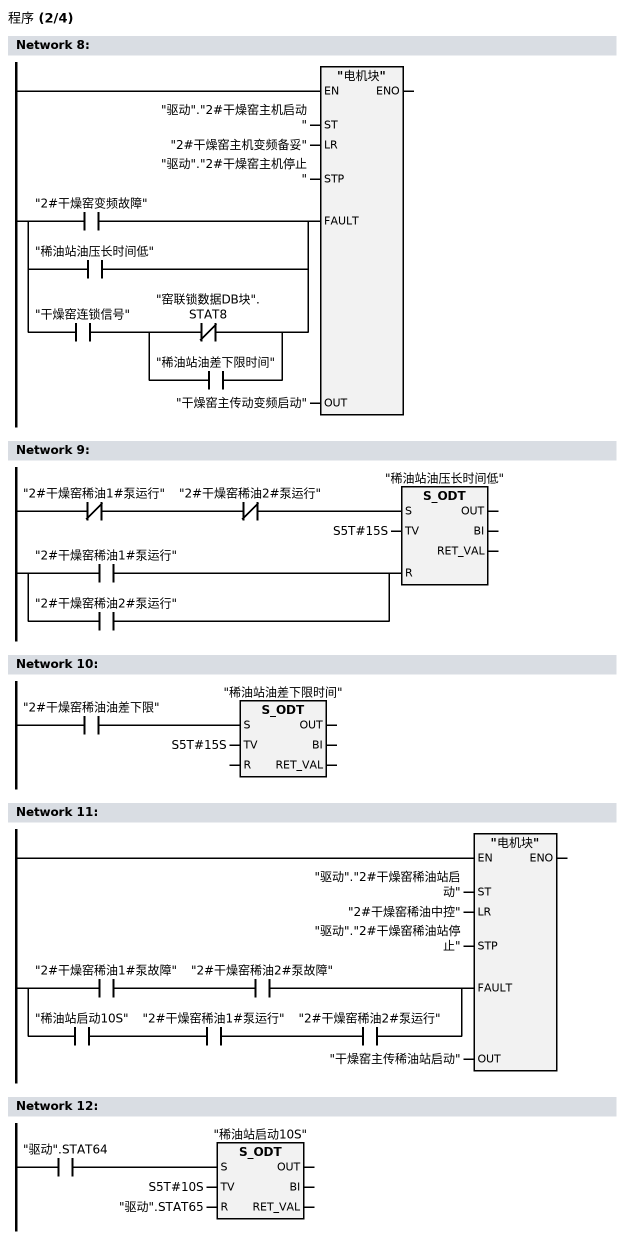
   RUNG wire#powerrail
      "电机块"(FAULT := wire#w2, ST := "驱动"."2#干燥窑主机启动", LR := "2#干燥窑主机变频备妥", STP := "驱动"."2#干燥窑主机停止", OUT := "干燥窑主传动变频启动")
   END_RUNG
   RUNG wire#powerrail
      Contact( "2#干燥窑变频故障" )
   END_RUNG wire#w2
   RUNG wire#powerrail
      Contact( "稀油站油压长时间低" )
   END_RUNG wire#w2
   RUNG wire#powerrail
      Contact( "干燥窑连锁信号" )
      wire#w1
      I_Contact( "窑联锁数据DB块".STAT8 )
   END_RUNG wire#w2
   RUNG wire#w1
      Contact( "稀油站油差下限时间" )
   END_RUNG wire#w2
   // the same network as SCL:
   "电机块"(ST := "驱动"."2#干燥窑主机启动",
         LR := "2#干燥窑主机变频备妥",
         STP := "驱动"."2#干燥窑主机停止",
         FAULT := "2#干燥窑变频故障" OR "稀油站油压长时间低" OR ("干燥窑连锁信号" AND (NOT "窑联锁数据DB块".STAT8 OR "稀油站油差下限时间")),
         OUT := "干燥窑主传动变频启动");
END_REGION

REGION Network 9
   RUNG wire#powerrail
      I_Contact( "2#干燥窑稀油1#泵运行" )
      I_Contact( "2#干燥窑稀油2#泵运行" )
      S_ODT(T_NO := "稀油站油压长时间低", TV := S5T#15S, R := wire#w1, BI =>, RET_VAL =>)
   END_RUNG
   RUNG wire#powerrail
      Contact( "2#干燥窑稀油1#泵运行" )
   END_RUNG wire#w1
   RUNG wire#powerrail
      Contact( "2#干燥窑稀油2#泵运行" )
   END_RUNG wire#w1
   // the same network as SCL:
   #_s5time1 := S_ODT(T_NO := "稀油站油压长时间低",
                      TV := S5T#15S,
                      R := "2#干燥窑稀油1#泵运行" OR "2#干燥窑稀油2#泵运行",
                      S := NOT "2#干燥窑稀油1#泵运行" AND NOT "2#干燥窑稀油2#泵运行");
END_REGION

REGION Network 10
   RUNG wire#powerrail
      Contact( "2#干燥窑稀油油差下限" )
      S_ODT(T_NO := "稀油站油差下限时间", TV := S5T#15S, R :=, BI =>, RET_VAL =>)
   END_RUNG
   // the same network as SCL:
   #_s5time1 := S_ODT(T_NO := "稀油站油差下限时间", TV := S5T#15S, S := "2#干燥窑稀油油差下限");
END_REGION

REGION Network 11
   RUNG wire#powerrail
      "电机块"(FAULT := wire#w1, ST := "驱动"."2#干燥窑稀油站启动", LR := "2#干燥窑稀油中控", STP := "驱动"."2#干燥窑稀油站停止", OUT := "干燥窑主传稀油站启动")
   END_RUNG
   RUNG wire#powerrail
      Contact( "2#干燥窑稀油1#泵故障" )
      Contact( "2#干燥窑稀油2#泵故障" )
   END_RUNG wire#w1
   RUNG wire#powerrail
      Contact( "稀油站启动10S" )
      Contact( "2#干燥窑稀油1#泵运行" )
      Contact( "2#干燥窑稀油2#泵运行" )
   END_RUNG wire#w1
   // the same network as SCL:
   "电机块"(ST := "驱动"."2#干燥窑稀油站启动",
         LR := "2#干燥窑稀油中控",
         STP := "驱动"."2#干燥窑稀油站停止",
         FAULT := ("2#干燥窑稀油1#泵故障" AND "2#干燥窑稀油2#泵故障") OR ("稀油站启动10S" AND "2#干燥窑稀油1#泵运行" AND "2#干燥窑稀油2#泵运行"),
         OUT := "干燥窑主传稀油站启动");
END_REGION

REGION Network 12
   RUNG wire#powerrail
      Contact( "驱动".STAT64 )
      S_ODT(T_NO := "稀油站启动10S", TV := S5T#10S, R := "驱动".STAT65, BI =>, RET_VAL =>)
   END_RUNG
   // the same network as SCL:
   #_s5time1 := S_ODT(T_NO := "稀油站启动10S", S := "驱动".STAT64, TV := S5T#10S, R := "驱动".STAT65);
END_REGION

REGION Network 13
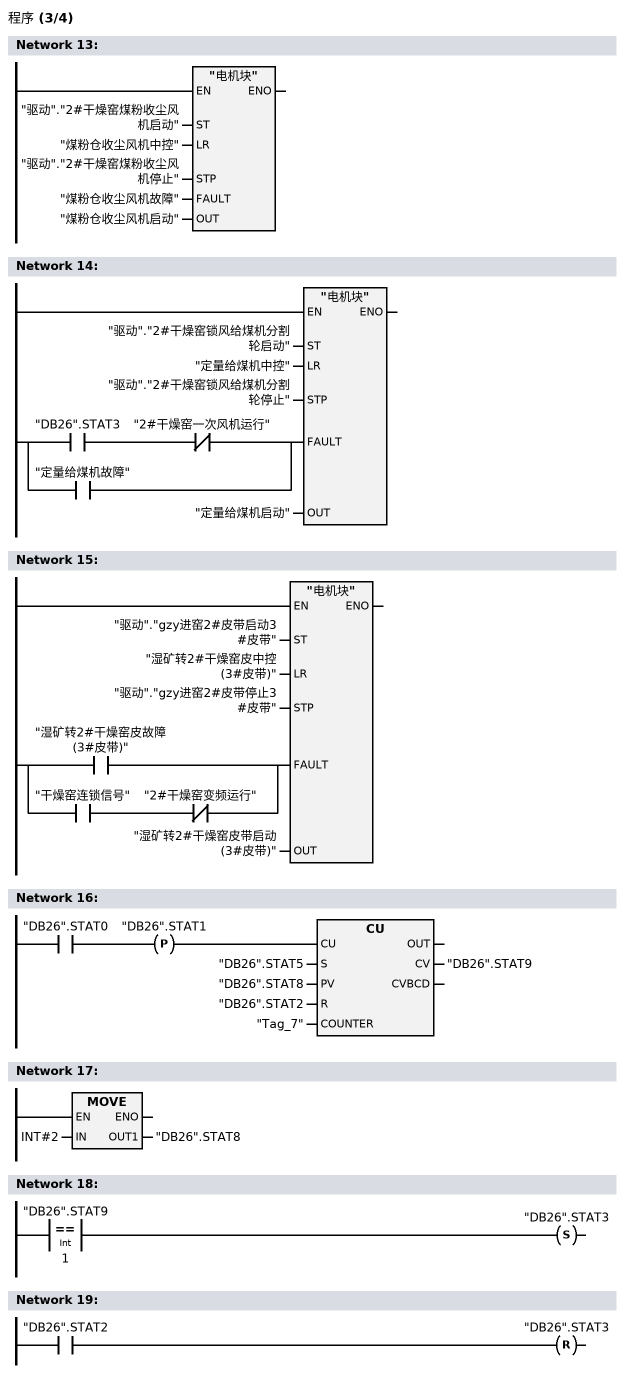
   RUNG wire#powerrail
      "电机块"(ST := "驱动"."2#干燥窑煤粉收尘风机启动", LR := "煤粉仓收尘风机中控", STP := "驱动"."2#干燥窑煤粉收尘风机停止", FAULT := "煤粉仓收尘风机故障", OUT := "煤粉仓收尘风机启动")
   END_RUNG
   // the same network as SCL:
   "电机块"(ST := "驱动"."2#干燥窑煤粉收尘风机启动",
         LR := "煤粉仓收尘风机中控",
         STP := "驱动"."2#干燥窑煤粉收尘风机停止",
         FAULT := "煤粉仓收尘风机故障",
         OUT := "煤粉仓收尘风机启动");
END_REGION

REGION Network 14
   RUNG wire#powerrail
      "电机块"(FAULT := wire#w1, ST := "驱动"."2#干燥窑锁风给煤机分割轮启动", LR := "定量给煤机中控", STP := "驱动"."2#干燥窑锁风给煤机分割轮停止", OUT := "定量给煤机启动")
   END_RUNG
   RUNG wire#powerrail
      Contact( "DB26".STAT3 )
      I_Contact( "2#干燥窑一次风机运行" )
   END_RUNG wire#w1
   RUNG wire#powerrail
      Contact( "定量给煤机故障" )
   END_RUNG wire#w1
   // the same network as SCL:
   "电机块"(ST := "驱动"."2#干燥窑锁风给煤机分割轮启动",
         LR := "定量给煤机中控",
         STP := "驱动"."2#干燥窑锁风给煤机分割轮停止",
         FAULT := ("DB26".STAT3 AND NOT "2#干燥窑一次风机运行") OR "定量给煤机故障",
         OUT := "定量给煤机启动");
END_REGION

REGION Network 15
   RUNG wire#powerrail
      "电机块"(FAULT := wire#w1, ST := "驱动"."gzy进窑2#皮带启动3#皮带", LR := "湿矿转2#干燥窑皮中控  (3#皮带)", STP := "驱动"."gzy进窑2#皮带停止3#皮带", OUT := "湿矿转2#干燥窑皮带启动  (3#皮带)")
   END_RUNG
   RUNG wire#powerrail
      Contact( "湿矿转2#干燥窑皮故障  (3#皮带)" )
   END_RUNG wire#w1
   RUNG wire#powerrail
      Contact( "干燥窑连锁信号" )
      I_Contact( "2#干燥窑变频运行" )
   END_RUNG wire#w1
   // the same network as SCL:
   "电机块"(ST := "驱动"."gzy进窑2#皮带启动3#皮带",
         LR := "湿矿转2#干燥窑皮中控  (3#皮带)",
         STP := "驱动"."gzy进窑2#皮带停止3#皮带",
         FAULT := "湿矿转2#干燥窑皮故障  (3#皮带)" OR ("干燥窑连锁信号" AND NOT "2#干燥窑变频运行"),
         OUT := "湿矿转2#干燥窑皮带启动  (3#皮带)");
END_REGION

REGION Network 16
   // no SCL statement known for Cu: written as a call
   #_w1 := "DB26".STAT0 AND NOT "DB26".STAT1;   // rising edge
   "DB26".STAT1 := "DB26".STAT0;
   Cu(cu := #_w1,
      s := "DB26".STAT5,
      pv := "DB26".STAT8,
      r := "DB26".STAT2,
      "counter" := "Tag_7",
      cv => "DB26".STAT9);
END_REGION

REGION Network 17
   RUNG wire#powerrail
      { S7_GenerateENO := "TRUE" } Move(in := INT#2, out1 => "DB26".STAT8)
   END_RUNG
   // the same network as SCL:
   "DB26".STAT8 := INT#2;
END_REGION

REGION Network 18
   RUNG wire#powerrail
      { S7_Templates := "SrcType := Int" } EQ_Contact(in1 := "DB26".STAT9, in2 := 1)
      S_Coil( "DB26".STAT3 )
   END_RUNG
   // the same network as SCL:
   IF "DB26".STAT9 = 1 THEN "DB26".STAT3 := TRUE; END_IF;
END_REGION

REGION Network 19
   RUNG wire#powerrail
      Contact( "DB26".STAT2 )
      R_Coil( "DB26".STAT3 )
   END_RUNG
   // the same network as SCL:
   IF "DB26".STAT2 THEN "DB26".STAT3 := FALSE; END_IF;
END_REGION

REGION Network 20
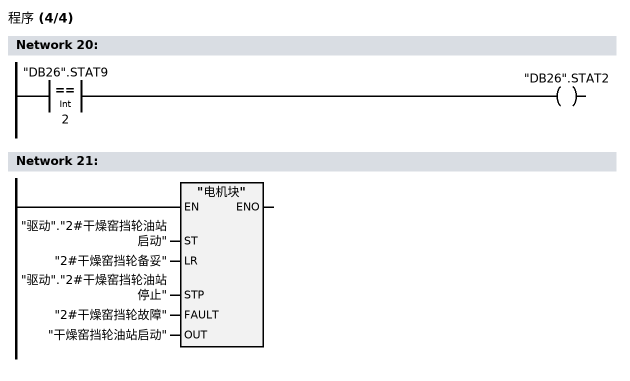
   RUNG wire#powerrail
      { S7_Templates := "SrcType := Int" } EQ_Contact(in1 := "DB26".STAT9, in2 := 2)
      Coil( "DB26".STAT2 )
   END_RUNG
   // the same network as SCL:
   "DB26".STAT2 := "DB26".STAT9 = 2;
END_REGION

REGION Network 21
   RUNG wire#powerrail
      "电机块"(ST := "驱动"."2#干燥窑挡轮油站启动", LR := "2#干燥窑挡轮备妥", STP := "驱动"."2#干燥窑挡轮油站停止", FAULT := "2#干燥窑挡轮故障", OUT := "干燥窑挡轮油站启动")
   END_RUNG
   // the same network as SCL:
   "电机块"(ST := "驱动"."2#干燥窑挡轮油站启动",
         LR := "2#干燥窑挡轮备妥",
         STP := "驱动"."2#干燥窑挡轮油站停止",
         FAULT := "2#干燥窑挡轮故障",
         OUT := "干燥窑挡轮油站启动");
END_REGION
END_FUNCTION

FUNCTION "FC4_粘料" : Void   // FC4, LAD
{ S7_Optimized_Access := 'TRUE' }
VERSION : 0.1
   VAR_TEMP   // added for the SCL form of the ladder/FBD networks
      _w1 : Bool;
      _w2 : Bool;
   END_VAR
BEGIN

REGION Network 1
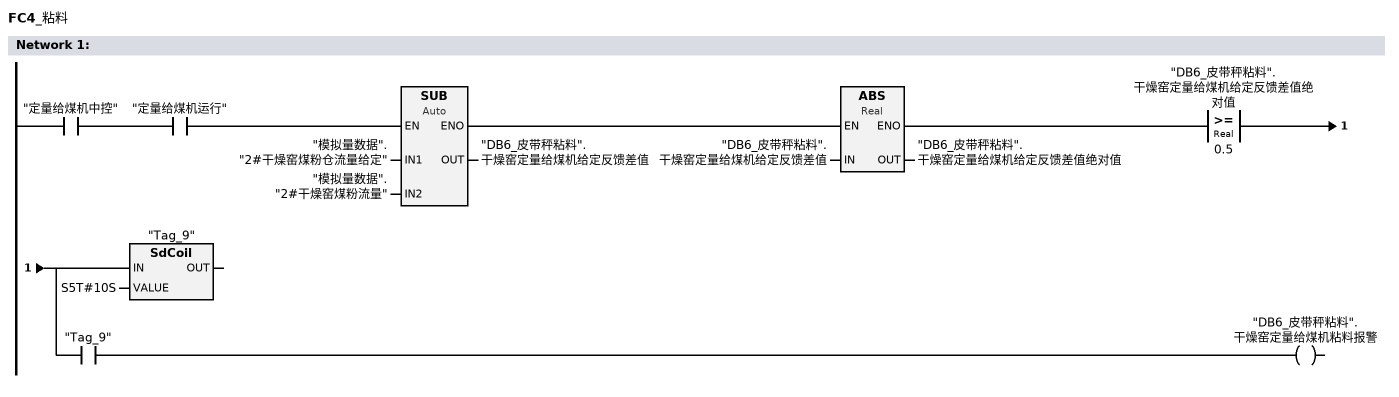
   // no SCL statement known for SdCoil: written as a call
   #_w1 := "定量给煤机中控" AND "定量给煤机运行";
   IF #_w1 THEN
       "DB6_皮带秤粘料".干燥窑定量给煤机给定反馈差值 := "模拟量数据"."2#干燥窑煤粉仓流量给定" - "模拟量数据"."2#干燥窑煤粉流量";
       "DB6_皮带秤粘料".干燥窑定量给煤机给定反馈差值绝对值 := ABS("DB6_皮带秤粘料".干燥窑定量给煤机给定反馈差值);
   END_IF;
   #_w2 := #_w1 AND ("DB6_皮带秤粘料".干燥窑定量给煤机给定反馈差值绝对值 >= 0.5);
   SdCoil(in := #_w2, value := S5T#10S, operand := "Tag_9");
   "DB6_皮带秤粘料".干燥窑定量给煤机粘料报警 := #_w2 AND "Tag_9";
END_REGION
END_FUNCTION

FUNCTION "澳泰温度巡检仪" : Void   // FC5, LAD
{ S7_Optimized_Access := 'FALSE' }
VERSION : 0.1
BEGIN

REGION Network 1
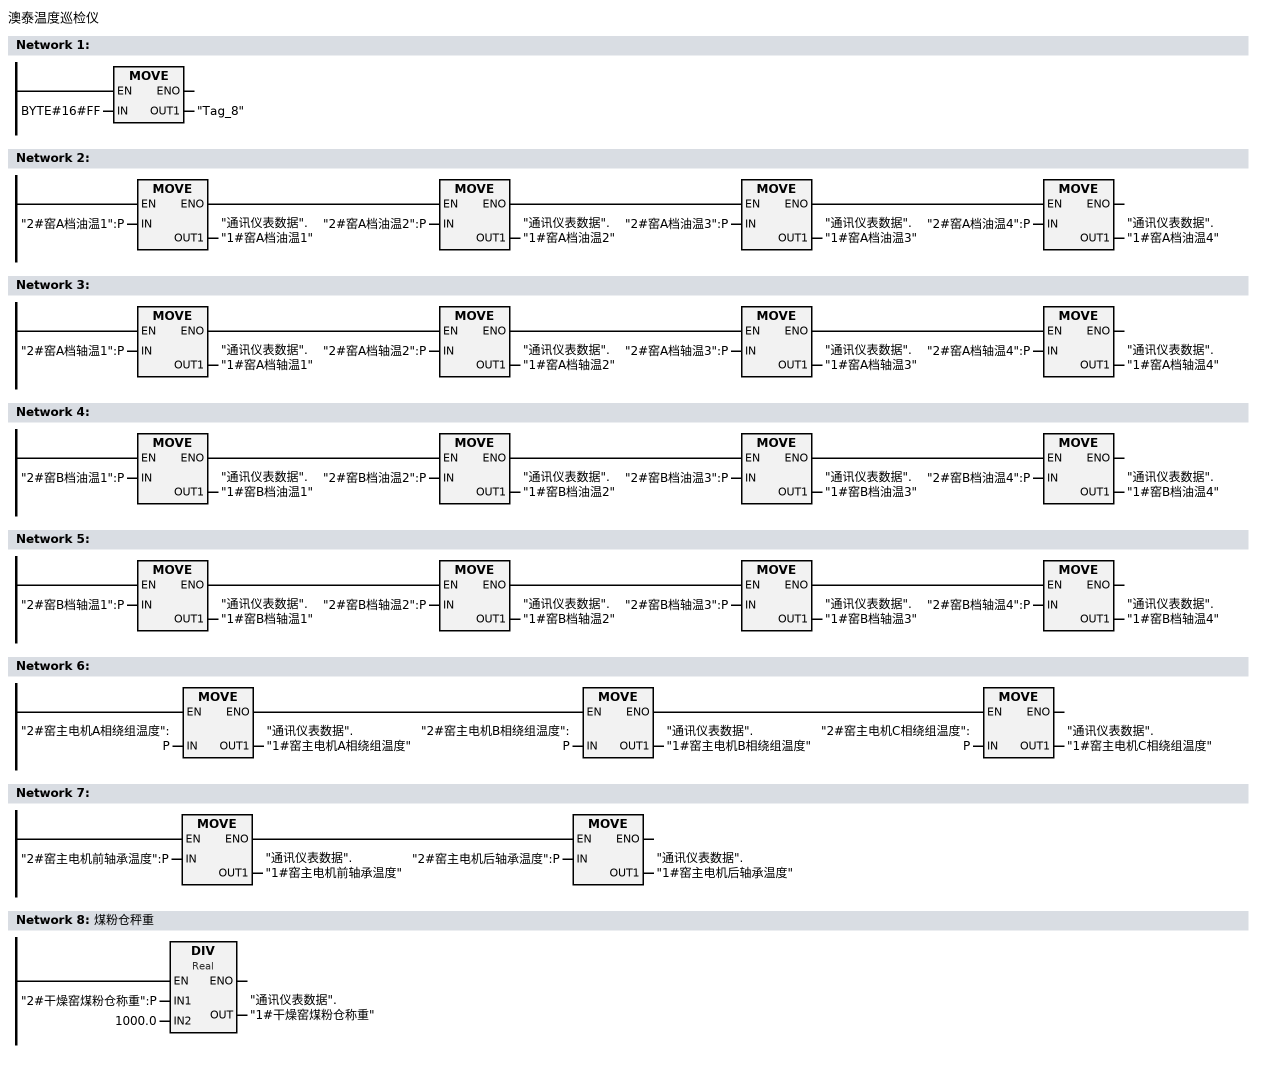
   RUNG wire#powerrail
      { S7_GenerateENO := "TRUE" } Move(in := BYTE#16#FF, out1 => "Tag_8")
   END_RUNG
   // the same network as SCL:
   "Tag_8" := BYTE#16#FF;
END_REGION

REGION Network 2
   RUNG wire#powerrail
      { S7_GenerateENO := "TRUE" } Move(in := "2#窑A档油温1":P, out1 => "通讯仪表数据"."1#窑A档油温1")
      { S7_GenerateENO := "TRUE" } Move(in := "2#窑A档油温2":P, out1 => "通讯仪表数据"."1#窑A档油温2")
      { S7_GenerateENO := "TRUE" } Move(in := "2#窑A档油温3":P, out1 => "通讯仪表数据"."1#窑A档油温3")
      { S7_GenerateENO := "TRUE" } Move(in := "2#窑A档油温4":P, out1 => "通讯仪表数据"."1#窑A档油温4")
   END_RUNG
   // the same network as SCL:
   // ENO of a box is taken as its EN; it also drops when the box reports an error
   "通讯仪表数据"."1#窑A档油温1" := "2#窑A档油温1":P;
   "通讯仪表数据"."1#窑A档油温2" := "2#窑A档油温2":P;
   "通讯仪表数据"."1#窑A档油温3" := "2#窑A档油温3":P;
   "通讯仪表数据"."1#窑A档油温4" := "2#窑A档油温4":P;
END_REGION

REGION Network 3
   RUNG wire#powerrail
      { S7_GenerateENO := "TRUE" } Move(in := "2#窑A档轴温1":P, out1 => "通讯仪表数据"."1#窑A档轴温1")
      { S7_GenerateENO := "TRUE" } Move(in := "2#窑A档轴温2":P, out1 => "通讯仪表数据"."1#窑A档轴温2")
      { S7_GenerateENO := "TRUE" } Move(in := "2#窑A档轴温3":P, out1 => "通讯仪表数据"."1#窑A档轴温3")
      { S7_GenerateENO := "TRUE" } Move(in := "2#窑A档轴温4":P, out1 => "通讯仪表数据"."1#窑A档轴温4")
   END_RUNG
   // the same network as SCL:
   // ENO of a box is taken as its EN; it also drops when the box reports an error
   "通讯仪表数据"."1#窑A档轴温1" := "2#窑A档轴温1":P;
   "通讯仪表数据"."1#窑A档轴温2" := "2#窑A档轴温2":P;
   "通讯仪表数据"."1#窑A档轴温3" := "2#窑A档轴温3":P;
   "通讯仪表数据"."1#窑A档轴温4" := "2#窑A档轴温4":P;
END_REGION

REGION Network 4
   RUNG wire#powerrail
      { S7_GenerateENO := "TRUE" } Move(in := "2#窑B档油温1":P, out1 => "通讯仪表数据"."1#窑B档油温1")
      { S7_GenerateENO := "TRUE" } Move(in := "2#窑B档油温2":P, out1 => "通讯仪表数据"."1#窑B档油温2")
      { S7_GenerateENO := "TRUE" } Move(in := "2#窑B档油温3":P, out1 => "通讯仪表数据"."1#窑B档油温3")
      { S7_GenerateENO := "TRUE" } Move(in := "2#窑B档油温4":P, out1 => "通讯仪表数据"."1#窑B档油温4")
   END_RUNG
   // the same network as SCL:
   // ENO of a box is taken as its EN; it also drops when the box reports an error
   "通讯仪表数据"."1#窑B档油温1" := "2#窑B档油温1":P;
   "通讯仪表数据"."1#窑B档油温2" := "2#窑B档油温2":P;
   "通讯仪表数据"."1#窑B档油温3" := "2#窑B档油温3":P;
   "通讯仪表数据"."1#窑B档油温4" := "2#窑B档油温4":P;
END_REGION

REGION Network 5
   RUNG wire#powerrail
      { S7_GenerateENO := "TRUE" } Move(in := "2#窑B档轴温1":P, out1 => "通讯仪表数据"."1#窑B档轴温1")
      { S7_GenerateENO := "TRUE" } Move(in := "2#窑B档轴温2":P, out1 => "通讯仪表数据"."1#窑B档轴温2")
      { S7_GenerateENO := "TRUE" } Move(in := "2#窑B档轴温3":P, out1 => "通讯仪表数据"."1#窑B档轴温3")
      { S7_GenerateENO := "TRUE" } Move(in := "2#窑B档轴温4":P, out1 => "通讯仪表数据"."1#窑B档轴温4")
   END_RUNG
   // the same network as SCL:
   // ENO of a box is taken as its EN; it also drops when the box reports an error
   "通讯仪表数据"."1#窑B档轴温1" := "2#窑B档轴温1":P;
   "通讯仪表数据"."1#窑B档轴温2" := "2#窑B档轴温2":P;
   "通讯仪表数据"."1#窑B档轴温3" := "2#窑B档轴温3":P;
   "通讯仪表数据"."1#窑B档轴温4" := "2#窑B档轴温4":P;
END_REGION

REGION Network 6
   RUNG wire#powerrail
      { S7_GenerateENO := "TRUE" } Move(in := "2#窑主电机A相绕组温度":P, out1 => "通讯仪表数据"."1#窑主电机A相绕组温度")
      { S7_GenerateENO := "TRUE" } Move(in := "2#窑主电机B相绕组温度":P, out1 => "通讯仪表数据"."1#窑主电机B相绕组温度")
      { S7_GenerateENO := "TRUE" } Move(in := "2#窑主电机C相绕组温度":P, out1 => "通讯仪表数据"."1#窑主电机C相绕组温度")
   END_RUNG
   // the same network as SCL:
   // ENO of a box is taken as its EN; it also drops when the box reports an error
   "通讯仪表数据"."1#窑主电机A相绕组温度" := "2#窑主电机A相绕组温度":P;
   "通讯仪表数据"."1#窑主电机B相绕组温度" := "2#窑主电机B相绕组温度":P;
   "通讯仪表数据"."1#窑主电机C相绕组温度" := "2#窑主电机C相绕组温度":P;
END_REGION

REGION Network 7
   RUNG wire#powerrail
      { S7_GenerateENO := "TRUE" } Move(in := "2#窑主电机前轴承温度":P, out1 => "通讯仪表数据"."1#窑主电机前轴承温度")
      { S7_GenerateENO := "TRUE" } Move(in := "2#窑主电机后轴承温度":P, out1 => "通讯仪表数据"."1#窑主电机后轴承温度")
   END_RUNG
   // the same network as SCL:
   // ENO of a box is taken as its EN; it also drops when the box reports an error
   "通讯仪表数据"."1#窑主电机前轴承温度" := "2#窑主电机前轴承温度":P;
   "通讯仪表数据"."1#窑主电机后轴承温度" := "2#窑主电机后轴承温度":P;
END_REGION

REGION Network 8: 煤粉仓秤重
   RUNG wire#powerrail
      { S7_Templates := "SrcType := Real" } Div(in1 := "2#干燥窑煤粉仓称重":P, in2 := 1000.0, out => "通讯仪表数据"."1#干燥窑煤粉仓称重")
   END_RUNG
   // the same network as SCL:
   "通讯仪表数据"."1#干燥窑煤粉仓称重" := "2#干燥窑煤粉仓称重":P / 1000.0;
END_REGION
END_FUNCTION

FUNCTION "1#2#干燥窑皮带联锁信号通" : Void   // FC16, LAD
{ S7_Optimized_Access := 'FALSE' }
VERSION : 0.1
BEGIN

REGION Network 1
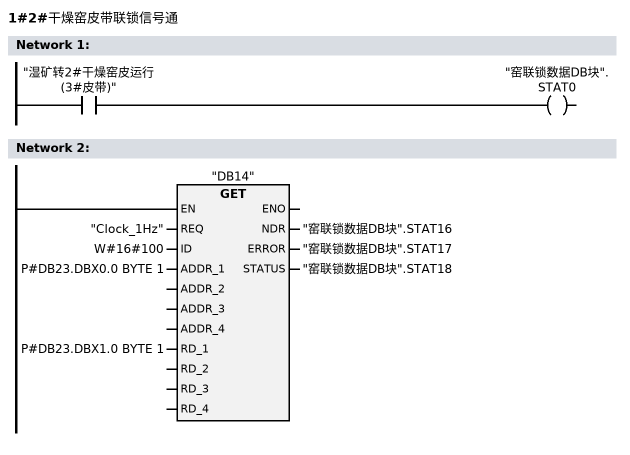
   RUNG wire#powerrail
      Contact( "湿矿转2#干燥窑皮运行  (3#皮带)" )
      Coil( "窑联锁数据DB块".STAT0 )
   END_RUNG
   // the same network as SCL:
   "窑联锁数据DB块".STAT0 := "湿矿转2#干燥窑皮运行  (3#皮带)";
END_REGION

REGION Network 2
   "DB14"(REQ := "Clock_1Hz",   // GET
          ID := W#16#100,
          ADDR_1 := P#DB23.DBX0.0 BYTE 1,
          RD_1 := P#DB23.DBX1.0 BYTE 1,
          NDR => "窑联锁数据DB块".STAT16,
          ERROR => "窑联锁数据DB块".STAT17,
          STATUS => "窑联锁数据DB块".STAT18);
END_REGION
END_FUNCTION

FUNCTION "模拟量转换" : Void   // FC21, LAD
{ S7_Optimized_Access := 'FALSE' }
VERSION : 0.1
BEGIN

REGION Network 1
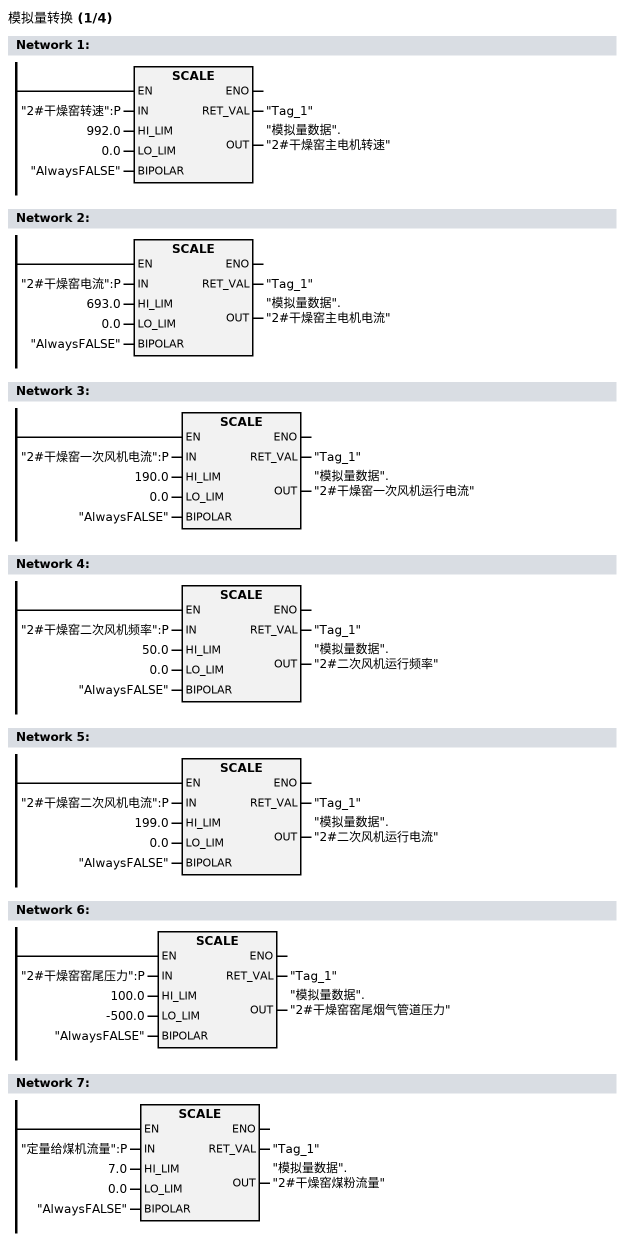
   "Tag_1" := SCALE(IN := "2#干燥窑转速":P,
                    HI_LIM := 992.0,
                    LO_LIM := 0.0,
                    BIPOLAR := "AlwaysFALSE",
                    OUT => "模拟量数据"."2#干燥窑主电机转速");
END_REGION

REGION Network 2
   "Tag_1" := SCALE(IN := "2#干燥窑电流":P,
                    HI_LIM := 693.0,
                    LO_LIM := 0.0,
                    BIPOLAR := "AlwaysFALSE",
                    OUT => "模拟量数据"."2#干燥窑主电机电流");
END_REGION

REGION Network 3
   "Tag_1" := SCALE(IN := "2#干燥窑一次风机电流":P,
                    HI_LIM := 190.0,
                    LO_LIM := 0.0,
                    BIPOLAR := "AlwaysFALSE",
                    OUT => "模拟量数据"."2#干燥窑一次风机运行电流");
END_REGION

REGION Network 4
   "Tag_1" := SCALE(IN := "2#干燥窑二次风机频率":P,
                    HI_LIM := 50.0,
                    LO_LIM := 0.0,
                    BIPOLAR := "AlwaysFALSE",
                    OUT => "模拟量数据"."2#二次风机运行频率");
END_REGION

REGION Network 5
   "Tag_1" := SCALE(IN := "2#干燥窑二次风机电流":P,
                    HI_LIM := 199.0,
                    LO_LIM := 0.0,
                    BIPOLAR := "AlwaysFALSE",
                    OUT => "模拟量数据"."2#二次风机运行电流");
END_REGION

REGION Network 6
   "Tag_1" := SCALE(IN := "2#干燥窑窑尾压力":P,
                    HI_LIM := 100.0,
                    LO_LIM := -500.0,
                    BIPOLAR := "AlwaysFALSE",
                    OUT => "模拟量数据"."2#干燥窑窑尾烟气管道压力");
END_REGION

REGION Network 7
   "Tag_1" := SCALE(IN := "定量给煤机流量":P,
                    HI_LIM := 7.0,
                    LO_LIM := 0.0,
                    BIPOLAR := "AlwaysFALSE",
                    OUT => "模拟量数据"."2#干燥窑煤粉流量");
END_REGION

REGION Network 8
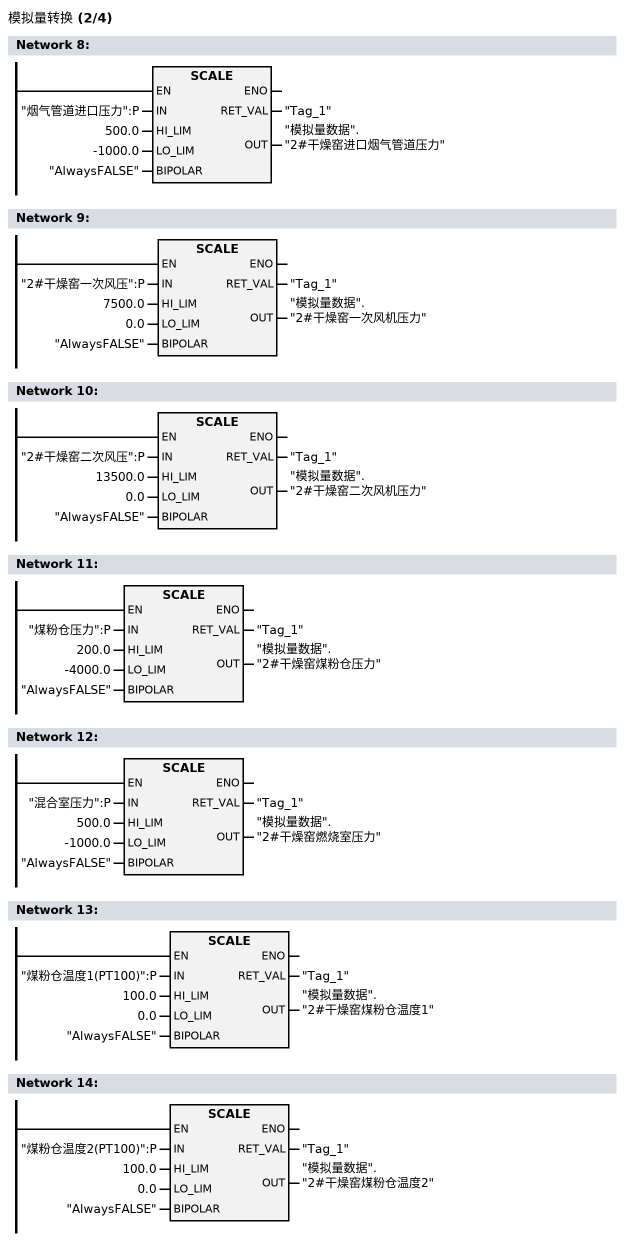
   "Tag_1" := SCALE(IN := "烟气管道进口压力":P,
                    HI_LIM := 500.0,
                    LO_LIM := -1000.0,
                    BIPOLAR := "AlwaysFALSE",
                    OUT => "模拟量数据"."2#干燥窑进口烟气管道压力");
END_REGION

REGION Network 9
   "Tag_1" := SCALE(IN := "2#干燥窑一次风压":P,
                    HI_LIM := 7500.0,
                    LO_LIM := 0.0,
                    BIPOLAR := "AlwaysFALSE",
                    OUT => "模拟量数据"."2#干燥窑一次风机压力");
END_REGION

REGION Network 10
   "Tag_1" := SCALE(IN := "2#干燥窑二次风压":P,
                    HI_LIM := 13500.0,
                    LO_LIM := 0.0,
                    BIPOLAR := "AlwaysFALSE",
                    OUT => "模拟量数据"."2#干燥窑二次风机压力");
END_REGION

REGION Network 11
   "Tag_1" := SCALE(IN := "煤粉仓压力":P,
                    HI_LIM := 200.0,
                    LO_LIM := -4000.0,
                    BIPOLAR := "AlwaysFALSE",
                    OUT => "模拟量数据"."2#干燥窑煤粉仓压力");
END_REGION

REGION Network 12
   "Tag_1" := SCALE(IN := "混合室压力":P,
                    HI_LIM := 500.0,
                    LO_LIM := -1000.0,
                    BIPOLAR := "AlwaysFALSE",
                    OUT => "模拟量数据"."2#干燥窑燃烧室压力");
END_REGION

REGION Network 13
   "Tag_1" := SCALE(IN := "煤粉仓温度1(PT100)":P,
                    HI_LIM := 100.0,
                    LO_LIM := 0.0,
                    BIPOLAR := "AlwaysFALSE",
                    OUT => "模拟量数据"."2#干燥窑煤粉仓温度1");
END_REGION

REGION Network 14
   "Tag_1" := SCALE(IN := "煤粉仓温度2(PT100)":P,
                    HI_LIM := 100.0,
                    LO_LIM := 0.0,
                    BIPOLAR := "AlwaysFALSE",
                    OUT => "模拟量数据"."2#干燥窑煤粉仓温度2");
END_REGION

REGION Network 15
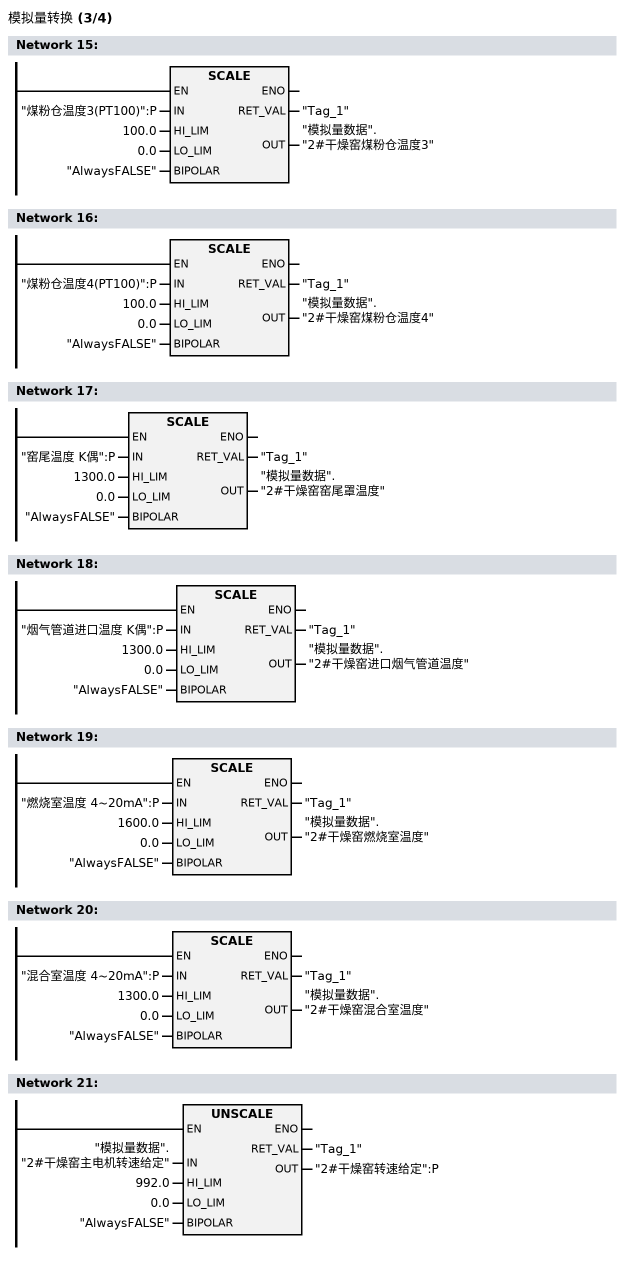
   "Tag_1" := SCALE(IN := "煤粉仓温度3(PT100)":P,
                    HI_LIM := 100.0,
                    LO_LIM := 0.0,
                    BIPOLAR := "AlwaysFALSE",
                    OUT => "模拟量数据"."2#干燥窑煤粉仓温度3");
END_REGION

REGION Network 16
   "Tag_1" := SCALE(IN := "煤粉仓温度4(PT100)":P,
                    HI_LIM := 100.0,
                    LO_LIM := 0.0,
                    BIPOLAR := "AlwaysFALSE",
                    OUT => "模拟量数据"."2#干燥窑煤粉仓温度4");
END_REGION

REGION Network 17
   "Tag_1" := SCALE(IN := "窑尾温度 K偶":P,
                    HI_LIM := 1300.0,
                    LO_LIM := 0.0,
                    BIPOLAR := "AlwaysFALSE",
                    OUT => "模拟量数据"."2#干燥窑窑尾罩温度");
END_REGION

REGION Network 18
   "Tag_1" := SCALE(IN := "烟气管道进口温度 K偶":P,
                    HI_LIM := 1300.0,
                    LO_LIM := 0.0,
                    BIPOLAR := "AlwaysFALSE",
                    OUT => "模拟量数据"."2#干燥窑进口烟气管道温度");
END_REGION

REGION Network 19
   "Tag_1" := SCALE(IN := "燃烧室温度 4~20mA":P,
                    HI_LIM := 1600.0,
                    LO_LIM := 0.0,
                    BIPOLAR := "AlwaysFALSE",
                    OUT => "模拟量数据"."2#干燥窑燃烧室温度");
END_REGION

REGION Network 20
   "Tag_1" := SCALE(IN := "混合室温度 4~20mA":P,
                    HI_LIM := 1300.0,
                    LO_LIM := 0.0,
                    BIPOLAR := "AlwaysFALSE",
                    OUT => "模拟量数据"."2#干燥窑混合室温度");
END_REGION

REGION Network 21
   "Tag_1" := UNSCALE(IN := "模拟量数据"."2#干燥窑主电机转速给定",
                      HI_LIM := 992.0,
                      LO_LIM := 0.0,
                      BIPOLAR := "AlwaysFALSE",
                      OUT => "2#干燥窑转速给定":P);
END_REGION

REGION Network 22
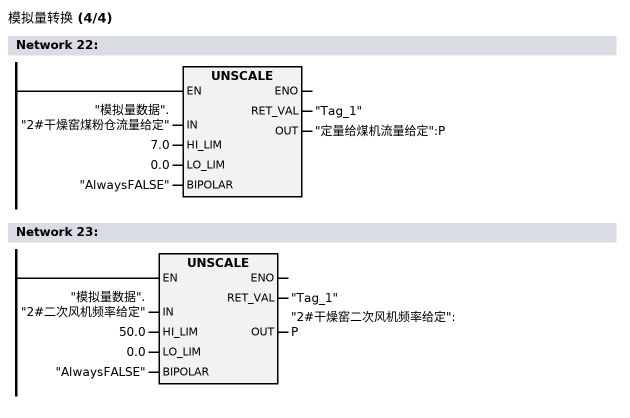
   "Tag_1" := UNSCALE(IN := "模拟量数据"."2#干燥窑煤粉仓流量给定",
                      HI_LIM := 7.0,
                      LO_LIM := 0.0,
                      BIPOLAR := "AlwaysFALSE",
                      OUT => "定量给煤机流量给定":P);
END_REGION

REGION Network 23
   "Tag_1" := UNSCALE(IN := "模拟量数据"."2#二次风机频率给定",
                      HI_LIM := 50.0,
                      LO_LIM := 0.0,
                      BIPOLAR := "AlwaysFALSE",
                      OUT => "2#干燥窑二次风机频率给定":P);
END_REGION
END_FUNCTION

FUNCTION "FC23" : Void   // FC23, LAD
{ S7_Optimized_Access := 'FALSE' }
VERSION : 0.1
   VAR_TEMP   // added for the SCL form of the ladder/FBD networks
      _w1 : Bool;
      _w2 : Bool;
   END_VAR
BEGIN

REGION Network 1
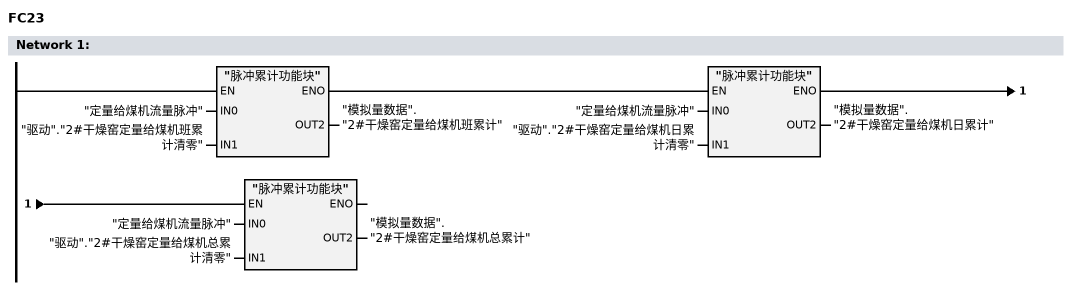
   RUNG wire#powerrail
      "脉冲累计功能块"(IN0 := "定量给煤机流量脉冲", IN1 := "驱动"."2#干燥窑定量给煤机班累计清零", OUT2 => "模拟量数据"."2#干燥窑定量给煤机班累计")
      "脉冲累计功能块"(IN0 := "定量给煤机流量脉冲", IN1 := "驱动"."2#干燥窑定量给煤机日累计清零", OUT2 => "模拟量数据"."2#干燥窑定量给煤机日累计")
      "脉冲累计功能块"(IN0 := "定量给煤机流量脉冲", IN1 := "驱动"."2#干燥窑定量给煤机总累计清零", OUT2 => "模拟量数据"."2#干燥窑定量给煤机总累计")
   END_RUNG
   // the same network as SCL:
   "脉冲累计功能块"(IN0 := "定量给煤机流量脉冲", IN1 := "驱动"."2#干燥窑定量给煤机班累计清零", OUT2 => "模拟量数据"."2#干燥窑定量给煤机班累计", ENO => #_w1);
   "脉冲累计功能块"(EN := #_w1,
             IN0 := "定量给煤机流量脉冲",
             IN1 := "驱动"."2#干燥窑定量给煤机日累计清零",
             OUT2 => "模拟量数据"."2#干燥窑定量给煤机日累计",
             ENO => #_w2);
   IF #_w2 THEN
       "脉冲累计功能块"(IN0 := "定量给煤机流量脉冲", IN1 := "驱动"."2#干燥窑定量给煤机总累计清零", OUT2 => "模拟量数据"."2#干燥窑定量给煤机总累计");
   END_IF;
END_REGION
END_FUNCTION

FUNCTION "FC40_DATA_ALARM" : Void   // FC40, LAD
{ S7_Optimized_Access := 'TRUE' }
VERSION : 0.1
BEGIN

REGION Network 1
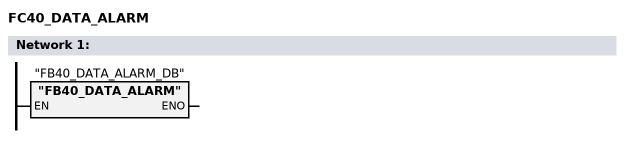
   RUNG wire#powerrail
      "FB40_DATA_ALARM_DB"()
   END_RUNG
   // the same network as SCL:
   "FB40_DATA_ALARM_DB"();   // "FB40_DATA_ALARM"
END_REGION
END_FUNCTION

FUNCTION "脉冲累计功能块" : Void   // FC116, LAD
{ S7_Optimized_Access := 'FALSE' }
VERSION : 0.1
   VAR_INPUT
      IN0 : Bool;
      IN1 : Bool;
   END_VAR
   VAR_OUTPUT
      OUT2 : Real;
   END_VAR
   VAR_TEMP
      TEMP3 : Bool;
      TEMP4 : Real;
      TEMP5 : Real;
      TEMP6 : Real;
   END_VAR
   VAR_TEMP   // added for the SCL form of the ladder/FBD networks
      _w1 : Bool;
   END_VAR
BEGIN

REGION Network 2